FUNCTION_BLOCK "1100_BWTS_CONTROL"   // FB1100, SCL
{ S7_Optimized_Access := 'TRUE' }
VERSION : 0.1
   VAR RETAIN
      State : "SYSTEM_STATES";   // Group of states required for BWT System
      TankData : Array[1..#NumberOfTanks] of "TANK_DATA";   // Group of tank data elements, one per tank on this system
   END_VAR
   VAR
      DECK_MANAGE_START_SUPPLY : "1110_DECK_MANAGE_START_SUPPLY";   // Function to start the deck supply (controlling CV valves 406, 407, 409, 411)
      DECK_MANAGE_STOP_SUPPLY : "1111_DECK_MANAGE_STOP_SUPPLY";   // Function to stop the deck supply (controlling CV valves 406, 407, 409, 411)
   END_VAR
   VAR RETAIN
      GTT_IN : "VALVE_GTT_IN";   // GTT Input data to management block
      GTT_OUT : "VALVE_GTT_OUT";   // GTT Output data from management block
      GTT_Exclusivity : "GTT_EXCLUSIVITY";   // GTT Exclusivity date to manage single valve actuation only
   END_VAR
   VAR
      GTT_MANAGE_VALVES : "1115_GTT_MANAGE_VALVES";
   END_VAR
   VAR RETAIN
      PVVX_IN : "VALVE_PVVX_IN";   // Vent A&B Input data to management blocks
      PVVX_OUT : "VALVE_PVVX_OUT";   // Vent A&B Output data from management blocks
   END_VAR
   VAR
      PVV_MANAGE_VALVES : "1120_PVV_MANAGE_VALVES";
      TANK_CONTROL_FPT : "1105_TANK_CONTROL";   // Tank sub-control block
      TANK_CONTROL_1P : "1105_TANK_CONTROL";   // Tank sub-control block
      TANK_CONTROL_1S : "1105_TANK_CONTROL";   // Tank sub-control block
      TANK_CONTROL_2P : "1105_TANK_CONTROL";   // Tank sub-control block
      TANK_CONTROL_2S : "1105_TANK_CONTROL";   // Tank sub-control block
      TANK_CONTROL_3P : "1105_TANK_CONTROL";   // Tank sub-control block
      TANK_CONTROL_3S : "1105_TANK_CONTROL";   // Tank sub-control block
      TANK_CONTROL_4P : "1105_TANK_CONTROL";   // Tank sub-control block
      TANK_CONTROL_4S : "1105_TANK_CONTROL";   // Tank sub-control block
      TANK_CONTROL_5P : "1105_TANK_CONTROL";   // Tank sub-control block
      TANK_CONTROL_5S : "1105_TANK_CONTROL";   // Tank sub-control block
      TANK_CONTROL_6P : "1105_TANK_CONTROL";   // Tank sub-control block
      TANK_CONTROL_6S : "1105_TANK_CONTROL";   // Tank sub-control block
      TANK_CONTROL_APT : "1105_TANK_CONTROL";   // Tank sub-control block
   END_VAR
   VAR RETAIN
      DWELL_TIMER : TONR_LTIME;   // Dwell Timer to manage Mid-Dwell period
      XEOX_TIMER : TONR_LTIME;   // DeOxygenation and ReOxygenation timer
      XEOX_PAUSE_TIMER : TONR_LTIME;   // The DeOxygenation Pause timer (with retain option)
      XEOX_PausedTime : LTime;   // A counter for the time spent in 'pause' whilst DeOxygenating.
      ShutdownStageReset : Bool := true;   // An reset flag for the shutdown procedure to set the stage to 0 once on a shutdown request.
   END_VAR
   VAR_TEMP
      Index : Int;   // Generic index for for loop parsing
      NextStageCheck : "ALARM_DEMAND_RTN";   // Temporary location for next stage alarm data and stage completion
      NextTreatmentGroup : Int;   // Temporary location for next treatment group calculation
   END_VAR
   VAR CONSTANT
      NumberOfTanks : Int := 14;   // Number of tanks in BWTS
      MaxTimerPT : LTime := LT#106751d;
      State_Init : Int := 0;   // State associated with State.System object.
      State_PreDwell : Int := 1;   // State associated with State.System object.
      State_DeOx : Int := 2;   // State associated with State.System object.
      State_DeOx_SupplyToDeck : Int := 200;   // Sate associated with State.DeOx object.
      State_DeOx_ClosePVV : Int := 201;   // Sate associated with State.DeOx object.
      State_DeOx_OpenGTT : Int := 202;   // Sate associated with State.DeOx object.
      State_DeOx_Monitor : Int := 203;   // Sate associated with State.DeOx object.
      State_DeOx_CloseGTT : Int := 204;   // Sate associated with State.DeOx object.
      State_DeOx_StopSupplyToDeck : Int := 205;   // Sate associated with State.DeOx object.
      State_DwellAndReOx : Int := 3;   // State associated with State.System object.
      State_DwellAndReOx_WaitMidDwell : Int := 300;   // Sate associated with State.ReOx object.
      State_DwellAndReOx_SupplyToDeck : Int := 301;   // Sate associated with State.ReOx object.
      State_DwellAndReOx_OpenPVV : Int := 302;   // Sate associated with State.ReOx object.
      State_DwellAndReOx_OpenGTT : Int := 303;   // Sate associated with State.ReOx object.
      State_DwellAndReOx_Monitor : Int := 304;   // Sate associated with State.ReOx object.
      State_DwellAndReOx_CloseGTT : Int := 305;   // Sate associated with State.ReOx object.
      State_DwellAndReOx_StopSupplyToDeck : Int := 306;   // Sate associated with State.ReOx object.
      State_DwellAndComplete : Int := 4;   // State associated with State.System object.
      State_DwellAndComplete_WaitPostDwell : Int := 400;   // Sate associated with State.Complete object.
      State_DwellAndComplete_Done : Int := 401;   // Sate associated with State.Complete object.
      State_Shutdown : Int := 5;   // State associated with State.System object.
      TankState_Init : Int := 1000;   // State associated with tank sub-control.
      TankState_PreDwell : Int := 1001;   // State associated with tank sub-control.
      TankState_DeOx : Int := 1002;   // State associated with tank sub-control.
      TankState_MidDwell : Int := 1003;   // State associated with tank sub-control.
      TankState_ReOx : Int := 1004;   // State associated with tank sub-control.
      TankState_PostDwell : Int := 1005;   // State associated with tank sub-control.
      TankState_Done : Int := 1006;   // State associated with tank sub-control.
   END_VAR
   // TankData[1].AllocatedTreatmentGroup := 1;
   // TankData[2].AllocatedTreatmentGroup := 1;
   // TankData[3].AllocatedTreatmentGroup := 1;
   // TankData[4].AllocatedTreatmentGroup := 2;
   // TankData[5].AllocatedTreatmentGroup := 2;
   // TankData[6].AllocatedTreatmentGroup := 2;
   // TankData[7].AllocatedTreatmentGroup := 2;
   // TankData[8].AllocatedTreatmentGroup := 3;
   // TankData[9].AllocatedTreatmentGroup := 3;
   // TankData[10].AllocatedTreatmentGroup := 3;
   // TankData[11].AllocatedTreatmentGroup := 4;
   // TankData[12].AllocatedTreatmentGroup := 4;
   // TankData[13].AllocatedTreatmentGroup := 4;
   // TankData[14].AllocatedTreatmentGroup := 4;
   // TankData[1].Active := False;
   // TankData[1].XeOx_Complete := False;
   // TankData[1].Timer_Complete := False;
   // TankData[2].Active := False;
   // TankData[2].XeOx_Complete := False;
   // TankData[2].Timer_Complete := False;
   // TankData[3].Active := False;
   // TankData[3].XeOx_Complete := False;
   // TankData[3].Timer_Complete := False;
   // TankData[4].Active := False;
   // TankData[4].XeOx_Complete := False;
   // TankData[4].Timer_Complete := False;
   // TankData[5].Active := False;
   // TankData[5].XeOx_Complete := False;
   // TankData[5].Timer_Complete := False;
   // TankData[6].Active := False;
   // TankData[6].XeOx_Complete := False;
   // TankData[6].Timer_Complete := False;
   // TankData[7].Active := False;
   // TankData[7].XeOx_Complete := False;
   // TankData[7].Timer_Complete := False;
   // TankData[8].Active := False;
   // TankData[8].XeOx_Complete := False;
   // TankData[8].Timer_Complete := False;
   // TankData[9].Active := False;
   // TankData[9].XeOx_Complete := False;
   // TankData[9].Timer_Complete := False;
   // TankData[10].Active := False;
   // TankData[10].XeOx_Complete := False;
   // TankData[10].Timer_Complete := False;
   // TankData[11].Active := False;
   // TankData[11].XeOx_Complete := False;
   // TankData[11].Timer_Complete := False;
   // TankData[12].Active := False;
   // TankData[12].XeOx_Complete := False;
   // TankData[12].Timer_Complete := False;
   // TankData[13].Active := False;
   // TankData[13].XeOx_Complete := False;
   // TankData[13].Timer_Complete := False;
   // TankData[14].Active := False;
   // TankData[14].XeOx_Complete := False;
   // TankData[14].Timer_Complete := False;
   // DECK_MANAGE_START_SUPPLY.DNC_500CV406.DemandIn := False;
   // DECK_MANAGE_START_SUPPLY.DNC_500CV406.NO_Type := False;
   // DECK_MANAGE_START_SUPPLY.DNC_500CV406.NC_Type := False;
   // DECK_MANAGE_START_SUPPLY.DNC_500CV406.ValveOpenStatus := False;
   // DECK_MANAGE_START_SUPPLY.DNC_500CV406.ValveClsdStatus := False;
   // DECK_MANAGE_START_SUPPLY.DNC_500CV406.DemandOut := False;
   // DECK_MANAGE_START_SUPPLY.DNC_500CV406.DemandComplete := False;
   // DECK_MANAGE_START_SUPPLY.DNC_500CV406.Alarm := False;
   // DECK_MANAGE_START_SUPPLY.DNC_500CV406.Healthy := False;
   // DECK_MANAGE_START_SUPPLY.DNC_500CV406.Config_Error := False;
   // DECK_MANAGE_START_SUPPLY.DNC_500CV406.Sensor_Fault := False;
   // DECK_MANAGE_START_SUPPLY.DNC_500CV406.TRAVEL_TIME.IN := False;
   // DECK_MANAGE_START_SUPPLY.DNC_600CV407.DemandIn := False;
   // DECK_MANAGE_START_SUPPLY.DNC_600CV407.NO_Type := False;
   // DECK_MANAGE_START_SUPPLY.DNC_600CV407.NC_Type := False;
   // DECK_MANAGE_START_SUPPLY.DNC_600CV407.ValveOpenStatus := False;
   // DECK_MANAGE_START_SUPPLY.DNC_600CV407.ValveClsdStatus := False;
   // DECK_MANAGE_START_SUPPLY.DNC_600CV407.DemandOut := False;
   // DECK_MANAGE_START_SUPPLY.DNC_600CV407.DemandComplete := False;
   // DECK_MANAGE_START_SUPPLY.DNC_600CV407.Alarm := False;
   // DECK_MANAGE_START_SUPPLY.DNC_600CV407.Healthy := False;
   // DECK_MANAGE_START_SUPPLY.DNC_600CV407.Config_Error := False;
   // DECK_MANAGE_START_SUPPLY.DNC_600CV407.Sensor_Fault := False;
   // DECK_MANAGE_START_SUPPLY.DNC_600CV407.TRAVEL_TIME.IN := False;
   // DECK_MANAGE_START_SUPPLY.DNC_600CV411.DemandIn := False;
   // DECK_MANAGE_START_SUPPLY.DNC_600CV411.NO_Type := False;
   // DECK_MANAGE_START_SUPPLY.DNC_600CV411.NC_Type := False;
   // DECK_MANAGE_START_SUPPLY.DNC_600CV411.ValveOpenStatus := False;
   // DECK_MANAGE_START_SUPPLY.DNC_600CV411.ValveClsdStatus := False;
   // DECK_MANAGE_START_SUPPLY.DNC_600CV411.DemandOut := False;
   // DECK_MANAGE_START_SUPPLY.DNC_600CV411.DemandComplete := False;
   // DECK_MANAGE_START_SUPPLY.DNC_600CV411.Alarm := False;
   // DECK_MANAGE_START_SUPPLY.DNC_600CV411.Healthy := False;
   // DECK_MANAGE_START_SUPPLY.DNC_600CV411.Config_Error := False;
   // DECK_MANAGE_START_SUPPLY.DNC_600CV411.Sensor_Fault := False;
   // DECK_MANAGE_START_SUPPLY.DNC_600CV411.TRAVEL_TIME.IN := False;
   // DECK_MANAGE_START_SUPPLY.DNC_600CV409.DemandIn := False;
   // DECK_MANAGE_START_SUPPLY.DNC_600CV409.NO_Type := False;
   // DECK_MANAGE_START_SUPPLY.DNC_600CV409.NC_Type := False;
   // DECK_MANAGE_START_SUPPLY.DNC_600CV409.ValveOpenStatus := False;
   // DECK_MANAGE_START_SUPPLY.DNC_600CV409.ValveClsdStatus := False;
   // DECK_MANAGE_START_SUPPLY.DNC_600CV409.DemandOut := False;
   // DECK_MANAGE_START_SUPPLY.DNC_600CV409.DemandComplete := False;
   // DECK_MANAGE_START_SUPPLY.DNC_600CV409.Alarm := False;
   // DECK_MANAGE_START_SUPPLY.DNC_600CV409.Healthy := False;
   // DECK_MANAGE_START_SUPPLY.DNC_600CV409.Config_Error := False;
   // DECK_MANAGE_START_SUPPLY.DNC_600CV409.Sensor_Fault := False;
   // DECK_MANAGE_START_SUPPLY.DNC_600CV409.TRAVEL_TIME.IN := False;
   // DECK_MANAGE_START_SUPPLY.ShutdownDemand := False;
   // DECK_MANAGE_STOP_SUPPLY.DNC_500CV406.DemandIn := False;
   // DECK_MANAGE_STOP_SUPPLY.DNC_500CV406.NO_Type := False;
   // DECK_MANAGE_STOP_SUPPLY.DNC_500CV406.NC_Type := False;
   // DECK_MANAGE_STOP_SUPPLY.DNC_500CV406.ValveOpenStatus := False;
   // DECK_MANAGE_STOP_SUPPLY.DNC_500CV406.ValveClsdStatus := False;
   // DECK_MANAGE_STOP_SUPPLY.DNC_500CV406.DemandOut := False;
   // DECK_MANAGE_STOP_SUPPLY.DNC_500CV406.DemandComplete := False;
   // DECK_MANAGE_STOP_SUPPLY.DNC_500CV406.Alarm := False;
   // DECK_MANAGE_STOP_SUPPLY.DNC_500CV406.Healthy := False;
   // DECK_MANAGE_STOP_SUPPLY.DNC_500CV406.Config_Error := False;
   // DECK_MANAGE_STOP_SUPPLY.DNC_500CV406.Sensor_Fault := False;
   // DECK_MANAGE_STOP_SUPPLY.DNC_500CV406.TRAVEL_TIME.IN := False;
   // DECK_MANAGE_STOP_SUPPLY.DNC_600CV407.DemandIn := False;
   // DECK_MANAGE_STOP_SUPPLY.DNC_600CV407.NO_Type := False;
   // DECK_MANAGE_STOP_SUPPLY.DNC_600CV407.NC_Type := False;
   // DECK_MANAGE_STOP_SUPPLY.DNC_600CV407.ValveOpenStatus := False;
   // DECK_MANAGE_STOP_SUPPLY.DNC_600CV407.ValveClsdStatus := False;
   // DECK_MANAGE_STOP_SUPPLY.DNC_600CV407.DemandOut := False;
   // DECK_MANAGE_STOP_SUPPLY.DNC_600CV407.DemandComplete := False;
   // DECK_MANAGE_STOP_SUPPLY.DNC_600CV407.Alarm := False;
   // DECK_MANAGE_STOP_SUPPLY.DNC_600CV407.Healthy := False;
   // DECK_MANAGE_STOP_SUPPLY.DNC_600CV407.Config_Error := False;
   // DECK_MANAGE_STOP_SUPPLY.DNC_600CV407.Sensor_Fault := False;
   // DECK_MANAGE_STOP_SUPPLY.DNC_600CV407.TRAVEL_TIME.IN := False;
   // DECK_MANAGE_STOP_SUPPLY.DNC_600CV411.DemandIn := False;
   // DECK_MANAGE_STOP_SUPPLY.DNC_600CV411.NO_Type := False;
   // DECK_MANAGE_STOP_SUPPLY.DNC_600CV411.NC_Type := False;
   // DECK_MANAGE_STOP_SUPPLY.DNC_600CV411.ValveOpenStatus := False;
   // DECK_MANAGE_STOP_SUPPLY.DNC_600CV411.ValveClsdStatus := False;
   // DECK_MANAGE_STOP_SUPPLY.DNC_600CV411.DemandOut := False;
   // DECK_MANAGE_STOP_SUPPLY.DNC_600CV411.DemandComplete := False;
   // DECK_MANAGE_STOP_SUPPLY.DNC_600CV411.Alarm := False;
   // DECK_MANAGE_STOP_SUPPLY.DNC_600CV411.Healthy := False;
   // DECK_MANAGE_STOP_SUPPLY.DNC_600CV411.Config_Error := False;
   // DECK_MANAGE_STOP_SUPPLY.DNC_600CV411.Sensor_Fault := False;
   // DECK_MANAGE_STOP_SUPPLY.DNC_600CV411.TRAVEL_TIME.IN := False;
   // DECK_MANAGE_STOP_SUPPLY.DNC_600CV409.DemandIn := False;
   // DECK_MANAGE_STOP_SUPPLY.DNC_600CV409.NO_Type := False;
   // DECK_MANAGE_STOP_SUPPLY.DNC_600CV409.NC_Type := False;
   // DECK_MANAGE_STOP_SUPPLY.DNC_600CV409.ValveOpenStatus := False;
   // DECK_MANAGE_STOP_SUPPLY.DNC_600CV409.ValveClsdStatus := False;
   // DECK_MANAGE_STOP_SUPPLY.DNC_600CV409.DemandOut := False;
   // DECK_MANAGE_STOP_SUPPLY.DNC_600CV409.DemandComplete := False;
   // DECK_MANAGE_STOP_SUPPLY.DNC_600CV409.Alarm := False;
   // DECK_MANAGE_STOP_SUPPLY.DNC_600CV409.Healthy := False;
   // DECK_MANAGE_STOP_SUPPLY.DNC_600CV409.Config_Error := False;
   // DECK_MANAGE_STOP_SUPPLY.DNC_600CV409.Sensor_Fault := False;
   // DECK_MANAGE_STOP_SUPPLY.DNC_600CV409.TRAVEL_TIME.IN := False;
   // DECK_MANAGE_STOP_SUPPLY.TON_DELAY.IN := False;
   // DECK_MANAGE_STOP_SUPPLY.ShutdownDemand := False;
   // DECK_MANAGE_STOP_SUPPLY.StopDeckSupplyDone := False;
   // GTT_IN.GTT_Actuate[1] := False;
   // GTT_IN.GTT_Actuate[2] := False;
   // GTT_IN.GTT_Actuate[3] := False;
   // GTT_IN.GTT_Actuate[4] := False;
   // GTT_IN.GTT_Actuate[5] := False;
   // GTT_IN.GTT_Actuate[6] := False;
   // GTT_IN.GTT_Actuate[7] := False;
   // GTT_IN.GTT_Actuate[8] := False;
   // GTT_IN.GTT_Actuate[9] := False;
   // GTT_IN.GTT_Actuate[10] := False;
   // GTT_IN.GTT_Actuate[11] := False;
   // GTT_IN.GTT_Actuate[12] := False;
   // GTT_IN.GTT_Actuate[13] := False;
   // GTT_IN.GTT_Actuate[14] := False;
   // GTT_IN.GTT_ValveDemands[1] := False;
   // GTT_IN.GTT_ValveDemands[2] := False;
   // GTT_IN.GTT_ValveDemands[3] := False;
   // GTT_IN.GTT_ValveDemands[4] := False;
   // GTT_IN.GTT_ValveDemands[5] := False;
   // GTT_IN.GTT_ValveDemands[6] := False;
   // GTT_IN.GTT_ValveDemands[7] := False;
   // GTT_IN.GTT_ValveDemands[8] := False;
   // GTT_IN.GTT_ValveDemands[9] := False;
   // GTT_IN.GTT_ValveDemands[10] := False;
   // GTT_IN.GTT_ValveDemands[11] := False;
   // GTT_IN.GTT_ValveDemands[12] := False;
   // GTT_IN.GTT_ValveDemands[13] := False;
   // GTT_IN.GTT_ValveDemands[14] := False;
   // GTT_OUT.GTT_DemandsCompleted[1] := False;
   // GTT_OUT.GTT_DemandsCompleted[2] := False;
   // GTT_OUT.GTT_DemandsCompleted[3] := False;
   // GTT_OUT.GTT_DemandsCompleted[4] := False;
   // GTT_OUT.GTT_DemandsCompleted[5] := False;
   // GTT_OUT.GTT_DemandsCompleted[6] := False;
   // GTT_OUT.GTT_DemandsCompleted[7] := False;
   // GTT_OUT.GTT_DemandsCompleted[8] := False;
   // GTT_OUT.GTT_DemandsCompleted[9] := False;
   // GTT_OUT.GTT_DemandsCompleted[10] := False;
   // GTT_OUT.GTT_DemandsCompleted[11] := False;
   // GTT_OUT.GTT_DemandsCompleted[12] := False;
   // GTT_OUT.GTT_DemandsCompleted[13] := False;
   // GTT_OUT.GTT_DemandsCompleted[14] := False;
   // GTT_OUT.GTT_Alarms[1] := False;
   // GTT_OUT.GTT_Alarms[2] := False;
   // GTT_OUT.GTT_Alarms[3] := False;
   // GTT_OUT.GTT_Alarms[4] := False;
   // GTT_OUT.GTT_Alarms[5] := False;
   // GTT_OUT.GTT_Alarms[6] := False;
   // GTT_OUT.GTT_Alarms[7] := False;
   // GTT_OUT.GTT_Alarms[8] := False;
   // GTT_OUT.GTT_Alarms[9] := False;
   // GTT_OUT.GTT_Alarms[10] := False;
   // GTT_OUT.GTT_Alarms[11] := False;
   // GTT_OUT.GTT_Alarms[12] := False;
   // GTT_OUT.GTT_Alarms[13] := False;
   // GTT_OUT.GTT_Alarms[14] := False;
   // GTT_Exclusivity.Tank_Exclusivity := False;
   // GTT_MANAGE_VALVES.GTT_IN.GTT_Actuate[1] := False;
   // GTT_MANAGE_VALVES.GTT_IN.GTT_Actuate[2] := False;
   // GTT_MANAGE_VALVES.GTT_IN.GTT_Actuate[3] := False;
   // GTT_MANAGE_VALVES.GTT_IN.GTT_Actuate[4] := False;
   // GTT_MANAGE_VALVES.GTT_IN.GTT_Actuate[5] := False;
   // GTT_MANAGE_VALVES.GTT_IN.GTT_Actuate[6] := False;
   // GTT_MANAGE_VALVES.GTT_IN.GTT_Actuate[7] := False;
   // GTT_MANAGE_VALVES.GTT_IN.GTT_Actuate[8] := False;
   // GTT_MANAGE_VALVES.GTT_IN.GTT_Actuate[9] := False;
   // GTT_MANAGE_VALVES.GTT_IN.GTT_Actuate[10] := False;
   // GTT_MANAGE_VALVES.GTT_IN.GTT_Actuate[11] := False;
   // GTT_MANAGE_VALVES.GTT_IN.GTT_Actuate[12] := False;
   // GTT_MANAGE_VALVES.GTT_IN.GTT_Actuate[13] := False;
   // GTT_MANAGE_VALVES.GTT_IN.GTT_Actuate[14] := False;
   // GTT_MANAGE_VALVES.GTT_IN.GTT_ValveDemands[1] := False;
   // GTT_MANAGE_VALVES.GTT_IN.GTT_ValveDemands[2] := False;
   // GTT_MANAGE_VALVES.GTT_IN.GTT_ValveDemands[3] := False;
   // GTT_MANAGE_VALVES.GTT_IN.GTT_ValveDemands[4] := False;
   // GTT_MANAGE_VALVES.GTT_IN.GTT_ValveDemands[5] := False;
   // GTT_MANAGE_VALVES.GTT_IN.GTT_ValveDemands[6] := False;
   // GTT_MANAGE_VALVES.GTT_IN.GTT_ValveDemands[7] := False;
   // GTT_MANAGE_VALVES.GTT_IN.GTT_ValveDemands[8] := False;
   // GTT_MANAGE_VALVES.GTT_IN.GTT_ValveDemands[9] := False;
   // GTT_MANAGE_VALVES.GTT_IN.GTT_ValveDemands[10] := False;
   // GTT_MANAGE_VALVES.GTT_IN.GTT_ValveDemands[11] := False;
   // GTT_MANAGE_VALVES.GTT_IN.GTT_ValveDemands[12] := False;
   // GTT_MANAGE_VALVES.GTT_IN.GTT_ValveDemands[13] := False;
   // GTT_MANAGE_VALVES.GTT_IN.GTT_ValveDemands[14] := False;
   // GTT_MANAGE_VALVES.DNC_FPT_GTT.DemandIn := False;
   // GTT_MANAGE_VALVES.DNC_FPT_GTT.NO_Type := False;
   // GTT_MANAGE_VALVES.DNC_FPT_GTT.NC_Type := False;
   // GTT_MANAGE_VALVES.DNC_FPT_GTT.ValveOpenStatus := False;
   // GTT_MANAGE_VALVES.DNC_FPT_GTT.ValveClsdStatus := False;
   // GTT_MANAGE_VALVES.DNC_FPT_GTT.DemandOut := False;
   // GTT_MANAGE_VALVES.DNC_FPT_GTT.DemandComplete := False;
   // GTT_MANAGE_VALVES.DNC_FPT_GTT.Alarm := False;
   // GTT_MANAGE_VALVES.DNC_FPT_GTT.Healthy := False;
   // GTT_MANAGE_VALVES.DNC_FPT_GTT.Config_Error := False;
   // GTT_MANAGE_VALVES.DNC_FPT_GTT.Sensor_Fault := False;
   // GTT_MANAGE_VALVES.DNC_FPT_GTT.TRAVEL_TIME.IN := False;
   // GTT_MANAGE_VALVES.DNC_1P_GTT.DemandIn := False;
   // GTT_MANAGE_VALVES.DNC_1P_GTT.NO_Type := False;
   // GTT_MANAGE_VALVES.DNC_1P_GTT.NC_Type := False;
   // GTT_MANAGE_VALVES.DNC_1P_GTT.ValveOpenStatus := False;
   // GTT_MANAGE_VALVES.DNC_1P_GTT.ValveClsdStatus := False;
   // GTT_MANAGE_VALVES.DNC_1P_GTT.DemandOut := False;
   // GTT_MANAGE_VALVES.DNC_1P_GTT.DemandComplete := False;
   // GTT_MANAGE_VALVES.DNC_1P_GTT.Alarm := False;
   // GTT_MANAGE_VALVES.DNC_1P_GTT.Healthy := False;
   // GTT_MANAGE_VALVES.DNC_1P_GTT.Config_Error := False;
   // GTT_MANAGE_VALVES.DNC_1P_GTT.Sensor_Fault := False;
   // GTT_MANAGE_VALVES.DNC_1P_GTT.TRAVEL_TIME.IN := False;
   // GTT_MANAGE_VALVES.DNC_1S_GTT.DemandIn := False;
   // GTT_MANAGE_VALVES.DNC_1S_GTT.NO_Type := False;
   // GTT_MANAGE_VALVES.DNC_1S_GTT.NC_Type := False;
   // GTT_MANAGE_VALVES.DNC_1S_GTT.ValveOpenStatus := False;
   // GTT_MANAGE_VALVES.DNC_1S_GTT.ValveClsdStatus := False;
   // GTT_MANAGE_VALVES.DNC_1S_GTT.DemandOut := False;
   // GTT_MANAGE_VALVES.DNC_1S_GTT.DemandComplete := False;
   // GTT_MANAGE_VALVES.DNC_1S_GTT.Alarm := False;
   // GTT_MANAGE_VALVES.DNC_1S_GTT.Healthy := False;
   // GTT_MANAGE_VALVES.DNC_1S_GTT.Config_Error := False;
   // GTT_MANAGE_VALVES.DNC_1S_GTT.Sensor_Fault := False;
   // GTT_MANAGE_VALVES.DNC_1S_GTT.TRAVEL_TIME.IN := False;
   // GTT_MANAGE_VALVES.DNC_2P_GTT.DemandIn := False;
   // GTT_MANAGE_VALVES.DNC_2P_GTT.NO_Type := False;
   // GTT_MANAGE_VALVES.DNC_2P_GTT.NC_Type := False;
   // GTT_MANAGE_VALVES.DNC_2P_GTT.ValveOpenStatus := False;
   // GTT_MANAGE_VALVES.DNC_2P_GTT.ValveClsdStatus := False;
   // GTT_MANAGE_VALVES.DNC_2P_GTT.DemandOut := False;
   // GTT_MANAGE_VALVES.DNC_2P_GTT.DemandComplete := False;
   // GTT_MANAGE_VALVES.DNC_2P_GTT.Alarm := False;
   // GTT_MANAGE_VALVES.DNC_2P_GTT.Healthy := False;
   // GTT_MANAGE_VALVES.DNC_2P_GTT.Config_Error := False;
   // GTT_MANAGE_VALVES.DNC_2P_GTT.Sensor_Fault := False;
   // GTT_MANAGE_VALVES.DNC_2P_GTT.TRAVEL_TIME.IN := False;
   // GTT_MANAGE_VALVES.DNC_2S_GTT.DemandIn := False;
   // GTT_MANAGE_VALVES.DNC_2S_GTT.NO_Type := False;
   // GTT_MANAGE_VALVES.DNC_2S_GTT.NC_Type := False;
   // GTT_MANAGE_VALVES.DNC_2S_GTT.ValveOpenStatus := False;
   // GTT_MANAGE_VALVES.DNC_2S_GTT.ValveClsdStatus := False;
   // GTT_MANAGE_VALVES.DNC_2S_GTT.DemandOut := False;
   // GTT_MANAGE_VALVES.DNC_2S_GTT.DemandComplete := False;
   // GTT_MANAGE_VALVES.DNC_2S_GTT.Alarm := False;
   // GTT_MANAGE_VALVES.DNC_2S_GTT.Healthy := False;
   // GTT_MANAGE_VALVES.DNC_2S_GTT.Config_Error := False;
   // GTT_MANAGE_VALVES.DNC_2S_GTT.Sensor_Fault := False;
   // GTT_MANAGE_VALVES.DNC_2S_GTT.TRAVEL_TIME.IN := False;
   // GTT_MANAGE_VALVES.DNC_3P_GTT.DemandIn := False;
   // GTT_MANAGE_VALVES.DNC_3P_GTT.NO_Type := False;
   // GTT_MANAGE_VALVES.DNC_3P_GTT.NC_Type := False;
   // GTT_MANAGE_VALVES.DNC_3P_GTT.ValveOpenStatus := False;
   // GTT_MANAGE_VALVES.DNC_3P_GTT.ValveClsdStatus := False;
   // GTT_MANAGE_VALVES.DNC_3P_GTT.DemandOut := False;
   // GTT_MANAGE_VALVES.DNC_3P_GTT.DemandComplete := False;
   // GTT_MANAGE_VALVES.DNC_3P_GTT.Alarm := False;
   // GTT_MANAGE_VALVES.DNC_3P_GTT.Healthy := False;
   // GTT_MANAGE_VALVES.DNC_3P_GTT.Config_Error := False;
   // GTT_MANAGE_VALVES.DNC_3P_GTT.Sensor_Fault := False;
   // GTT_MANAGE_VALVES.DNC_3P_GTT.TRAVEL_TIME.IN := False;
   // GTT_MANAGE_VALVES.DNC_3S_GTT.DemandIn := False;
   // GTT_MANAGE_VALVES.DNC_3S_GTT.NO_Type := False;
   // GTT_MANAGE_VALVES.DNC_3S_GTT.NC_Type := False;
   // GTT_MANAGE_VALVES.DNC_3S_GTT.ValveOpenStatus := False;
   // GTT_MANAGE_VALVES.DNC_3S_GTT.ValveClsdStatus := False;
   // GTT_MANAGE_VALVES.DNC_3S_GTT.DemandOut := False;
   // GTT_MANAGE_VALVES.DNC_3S_GTT.DemandComplete := False;
   // GTT_MANAGE_VALVES.DNC_3S_GTT.Alarm := False;
   // GTT_MANAGE_VALVES.DNC_3S_GTT.Healthy := False;
   // GTT_MANAGE_VALVES.DNC_3S_GTT.Config_Error := False;
   // GTT_MANAGE_VALVES.DNC_3S_GTT.Sensor_Fault := False;
   // GTT_MANAGE_VALVES.DNC_3S_GTT.TRAVEL_TIME.IN := False;
   // GTT_MANAGE_VALVES.DNC_4P_GTT.DemandIn := False;
   // GTT_MANAGE_VALVES.DNC_4P_GTT.NO_Type := False;
   // GTT_MANAGE_VALVES.DNC_4P_GTT.NC_Type := False;
   // GTT_MANAGE_VALVES.DNC_4P_GTT.ValveOpenStatus := False;
   // GTT_MANAGE_VALVES.DNC_4P_GTT.ValveClsdStatus := False;
   // GTT_MANAGE_VALVES.DNC_4P_GTT.DemandOut := False;
   // GTT_MANAGE_VALVES.DNC_4P_GTT.DemandComplete := False;
   // GTT_MANAGE_VALVES.DNC_4P_GTT.Alarm := False;
   // GTT_MANAGE_VALVES.DNC_4P_GTT.Healthy := False;
   // GTT_MANAGE_VALVES.DNC_4P_GTT.Config_Error := False;
   // GTT_MANAGE_VALVES.DNC_4P_GTT.Sensor_Fault := False;
   // GTT_MANAGE_VALVES.DNC_4P_GTT.TRAVEL_TIME.IN := False;
   // GTT_MANAGE_VALVES.DNC_4S_GTT.DemandIn := False;
   // GTT_MANAGE_VALVES.DNC_4S_GTT.NO_Type := False;
   // GTT_MANAGE_VALVES.DNC_4S_GTT.NC_Type := False;
   // GTT_MANAGE_VALVES.DNC_4S_GTT.ValveOpenStatus := False;
   // GTT_MANAGE_VALVES.DNC_4S_GTT.ValveClsdStatus := False;
   // GTT_MANAGE_VALVES.DNC_4S_GTT.DemandOut := False;
   // GTT_MANAGE_VALVES.DNC_4S_GTT.DemandComplete := False;
   // GTT_MANAGE_VALVES.DNC_4S_GTT.Alarm := False;
   // GTT_MANAGE_VALVES.DNC_4S_GTT.Healthy := False;
   // GTT_MANAGE_VALVES.DNC_4S_GTT.Config_Error := False;
   // GTT_MANAGE_VALVES.DNC_4S_GTT.Sensor_Fault := False;
   // GTT_MANAGE_VALVES.DNC_4S_GTT.TRAVEL_TIME.IN := False;
   // GTT_MANAGE_VALVES.DNC_5P_GTT.DemandIn := False;
   // GTT_MANAGE_VALVES.DNC_5P_GTT.NO_Type := False;
   // GTT_MANAGE_VALVES.DNC_5P_GTT.NC_Type := False;
   // GTT_MANAGE_VALVES.DNC_5P_GTT.ValveOpenStatus := False;
   // GTT_MANAGE_VALVES.DNC_5P_GTT.ValveClsdStatus := False;
   // GTT_MANAGE_VALVES.DNC_5P_GTT.DemandOut := False;
   // GTT_MANAGE_VALVES.DNC_5P_GTT.DemandComplete := False;
   // GTT_MANAGE_VALVES.DNC_5P_GTT.Alarm := False;
   // GTT_MANAGE_VALVES.DNC_5P_GTT.Healthy := False;
   // GTT_MANAGE_VALVES.DNC_5P_GTT.Config_Error := False;
   // GTT_MANAGE_VALVES.DNC_5P_GTT.Sensor_Fault := False;
   // GTT_MANAGE_VALVES.DNC_5P_GTT.TRAVEL_TIME.IN := False;
   // GTT_MANAGE_VALVES.DNC_5S_GTT.DemandIn := False;
   // GTT_MANAGE_VALVES.DNC_5S_GTT.NO_Type := False;
   // GTT_MANAGE_VALVES.DNC_5S_GTT.NC_Type := False;
   // GTT_MANAGE_VALVES.DNC_5S_GTT.ValveOpenStatus := False;
   // GTT_MANAGE_VALVES.DNC_5S_GTT.ValveClsdStatus := False;
   // GTT_MANAGE_VALVES.DNC_5S_GTT.DemandOut := False;
   // GTT_MANAGE_VALVES.DNC_5S_GTT.DemandComplete := False;
   // GTT_MANAGE_VALVES.DNC_5S_GTT.Alarm := False;
   // GTT_MANAGE_VALVES.DNC_5S_GTT.Healthy := False;
   // GTT_MANAGE_VALVES.DNC_5S_GTT.Config_Error := False;
   // GTT_MANAGE_VALVES.DNC_5S_GTT.Sensor_Fault := False;
   // GTT_MANAGE_VALVES.DNC_5S_GTT.TRAVEL_TIME.IN := False;
   // GTT_MANAGE_VALVES.DNC_6P_GTT.DemandIn := False;
   // GTT_MANAGE_VALVES.DNC_6P_GTT.NO_Type := False;
   // GTT_MANAGE_VALVES.DNC_6P_GTT.NC_Type := False;
   // GTT_MANAGE_VALVES.DNC_6P_GTT.ValveOpenStatus := False;
   // GTT_MANAGE_VALVES.DNC_6P_GTT.ValveClsdStatus := False;
   // GTT_MANAGE_VALVES.DNC_6P_GTT.DemandOut := False;
   // GTT_MANAGE_VALVES.DNC_6P_GTT.DemandComplete := False;
   // GTT_MANAGE_VALVES.DNC_6P_GTT.Alarm := False;
   // GTT_MANAGE_VALVES.DNC_6P_GTT.Healthy := False;
   // GTT_MANAGE_VALVES.DNC_6P_GTT.Config_Error := False;
   // GTT_MANAGE_VALVES.DNC_6P_GTT.Sensor_Fault := False;
   // GTT_MANAGE_VALVES.DNC_6P_GTT.TRAVEL_TIME.IN := False;
   // GTT_MANAGE_VALVES.DNC_6S_GTT.DemandIn := False;
   // GTT_MANAGE_VALVES.DNC_6S_GTT.NO_Type := False;
   // GTT_MANAGE_VALVES.DNC_6S_GTT.NC_Type := False;
   // GTT_MANAGE_VALVES.DNC_6S_GTT.ValveOpenStatus := False;
   // GTT_MANAGE_VALVES.DNC_6S_GTT.ValveClsdStatus := False;
   // GTT_MANAGE_VALVES.DNC_6S_GTT.DemandOut := False;
   // GTT_MANAGE_VALVES.DNC_6S_GTT.DemandComplete := False;
   // GTT_MANAGE_VALVES.DNC_6S_GTT.Alarm := False;
   // GTT_MANAGE_VALVES.DNC_6S_GTT.Healthy := False;
   // GTT_MANAGE_VALVES.DNC_6S_GTT.Config_Error := False;
   // GTT_MANAGE_VALVES.DNC_6S_GTT.Sensor_Fault := False;
   // GTT_MANAGE_VALVES.DNC_6S_GTT.TRAVEL_TIME.IN := False;
   // GTT_MANAGE_VALVES.DNC_APT_GTT.DemandIn := False;
   // GTT_MANAGE_VALVES.DNC_APT_GTT.NO_Type := False;
   // GTT_MANAGE_VALVES.DNC_APT_GTT.NC_Type := False;
   // GTT_MANAGE_VALVES.DNC_APT_GTT.ValveOpenStatus := False;
   // GTT_MANAGE_VALVES.DNC_APT_GTT.ValveClsdStatus := False;
   // GTT_MANAGE_VALVES.DNC_APT_GTT.DemandOut := False;
   // GTT_MANAGE_VALVES.DNC_APT_GTT.DemandComplete := False;
   // GTT_MANAGE_VALVES.DNC_APT_GTT.Alarm := False;
   // GTT_MANAGE_VALVES.DNC_APT_GTT.Healthy := False;
   // GTT_MANAGE_VALVES.DNC_APT_GTT.Config_Error := False;
   // GTT_MANAGE_VALVES.DNC_APT_GTT.Sensor_Fault := False;
   // GTT_MANAGE_VALVES.DNC_APT_GTT.TRAVEL_TIME.IN := False;
   // PVVX_IN.PVVx_Actuate[1] := False;
   // PVVX_IN.PVVx_Actuate[2] := False;
   // PVVX_IN.PVVx_Actuate[3] := False;
   // PVVX_IN.PVVx_Actuate[4] := False;
   // PVVX_IN.PVVx_Actuate[5] := False;
   // PVVX_IN.PVVx_Actuate[6] := False;
   // PVVX_IN.PVVx_Actuate[7] := False;
   // PVVX_IN.PVVx_Actuate[8] := False;
   // PVVX_IN.PVVx_Actuate[9] := False;
   // PVVX_IN.PVVx_Actuate[10] := False;
   // PVVX_IN.PVVx_Actuate[11] := False;
   // PVVX_IN.PVVx_Actuate[12] := False;
   // PVVX_IN.PVVx_Actuate[13] := False;
   // PVVX_IN.PVVx_Actuate[14] := False;
   // PVVX_IN.PVVA_ValveDemands[1] := False;
   // PVVX_IN.PVVA_ValveDemands[2] := False;
   // PVVX_IN.PVVA_ValveDemands[3] := False;
   // PVVX_IN.PVVA_ValveDemands[4] := False;
   // PVVX_IN.PVVA_ValveDemands[5] := False;
   // PVVX_IN.PVVA_ValveDemands[6] := False;
   // PVVX_IN.PVVA_ValveDemands[7] := False;
   // PVVX_IN.PVVA_ValveDemands[8] := False;
   // PVVX_IN.PVVA_ValveDemands[9] := False;
   // PVVX_IN.PVVA_ValveDemands[10] := False;
   // PVVX_IN.PVVA_ValveDemands[11] := False;
   // PVVX_IN.PVVA_ValveDemands[12] := False;
   // PVVX_IN.PVVA_ValveDemands[13] := False;
   // PVVX_IN.PVVA_ValveDemands[14] := False;
   // PVVX_IN.PVVB_ValveDemands[1] := False;
   // PVVX_IN.PVVB_ValveDemands[2] := False;
   // PVVX_IN.PVVB_ValveDemands[3] := False;
   // PVVX_IN.PVVB_ValveDemands[4] := False;
   // PVVX_IN.PVVB_ValveDemands[5] := False;
   // PVVX_IN.PVVB_ValveDemands[6] := False;
   // PVVX_IN.PVVB_ValveDemands[7] := False;
   // PVVX_IN.PVVB_ValveDemands[8] := False;
   // PVVX_IN.PVVB_ValveDemands[9] := False;
   // PVVX_IN.PVVB_ValveDemands[10] := False;
   // PVVX_IN.PVVB_ValveDemands[11] := False;
   // PVVX_IN.PVVB_ValveDemands[12] := False;
   // PVVX_IN.PVVB_ValveDemands[13] := False;
   // PVVX_IN.PVVB_ValveDemands[14] := False;
   // PVVX_OUT.PVVA_DemandsCompleted[1] := False;
   // PVVX_OUT.PVVA_DemandsCompleted[2] := False;
   // PVVX_OUT.PVVA_DemandsCompleted[3] := False;
   // PVVX_OUT.PVVA_DemandsCompleted[4] := False;
   // PVVX_OUT.PVVA_DemandsCompleted[5] := False;
   // PVVX_OUT.PVVA_DemandsCompleted[6] := False;
   // PVVX_OUT.PVVA_DemandsCompleted[7] := False;
   // PVVX_OUT.PVVA_DemandsCompleted[8] := False;
   // PVVX_OUT.PVVA_DemandsCompleted[9] := False;
   // PVVX_OUT.PVVA_DemandsCompleted[10] := False;
   // PVVX_OUT.PVVA_DemandsCompleted[11] := False;
   // PVVX_OUT.PVVA_DemandsCompleted[12] := False;
   // PVVX_OUT.PVVA_DemandsCompleted[13] := False;
   // PVVX_OUT.PVVA_DemandsCompleted[14] := False;
   // PVVX_OUT.PVVA_Alarms[1] := False;
   // PVVX_OUT.PVVA_Alarms[2] := False;
   // PVVX_OUT.PVVA_Alarms[3] := False;
   // PVVX_OUT.PVVA_Alarms[4] := False;
   // PVVX_OUT.PVVA_Alarms[5] := False;
   // PVVX_OUT.PVVA_Alarms[6] := False;
   // PVVX_OUT.PVVA_Alarms[7] := False;
   // PVVX_OUT.PVVA_Alarms[8] := False;
   // PVVX_OUT.PVVA_Alarms[9] := False;
   // PVVX_OUT.PVVA_Alarms[10] := False;
   // PVVX_OUT.PVVA_Alarms[11] := False;
   // PVVX_OUT.PVVA_Alarms[12] := False;
   // PVVX_OUT.PVVA_Alarms[13] := False;
   // PVVX_OUT.PVVA_Alarms[14] := False;
   // PVVX_OUT.PVVB_DemandsCompleted[1] := False;
   // PVVX_OUT.PVVB_DemandsCompleted[2] := False;
   // PVVX_OUT.PVVB_DemandsCompleted[3] := False;
   // PVVX_OUT.PVVB_DemandsCompleted[4] := False;
   // PVVX_OUT.PVVB_DemandsCompleted[5] := False;
   // PVVX_OUT.PVVB_DemandsCompleted[6] := False;
   // PVVX_OUT.PVVB_DemandsCompleted[7] := False;
   // PVVX_OUT.PVVB_DemandsCompleted[8] := False;
   // PVVX_OUT.PVVB_DemandsCompleted[9] := False;
   // PVVX_OUT.PVVB_DemandsCompleted[10] := False;
   // PVVX_OUT.PVVB_DemandsCompleted[11] := False;
   // PVVX_OUT.PVVB_DemandsCompleted[12] := False;
   // PVVX_OUT.PVVB_DemandsCompleted[13] := False;
   // PVVX_OUT.PVVB_DemandsCompleted[14] := False;
   // PVVX_OUT.PVVB_Alarms[1] := False;
   // PVVX_OUT.PVVB_Alarms[2] := False;
   // PVVX_OUT.PVVB_Alarms[3] := False;
   // PVVX_OUT.PVVB_Alarms[4] := False;
   // PVVX_OUT.PVVB_Alarms[5] := False;
   // PVVX_OUT.PVVB_Alarms[6] := False;
   // PVVX_OUT.PVVB_Alarms[7] := False;
   // PVVX_OUT.PVVB_Alarms[8] := False;
   // PVVX_OUT.PVVB_Alarms[9] := False;
   // PVVX_OUT.PVVB_Alarms[10] := False;
   // PVVX_OUT.PVVB_Alarms[11] := False;
   // PVVX_OUT.PVVB_Alarms[12] := False;
   // PVVX_OUT.PVVB_Alarms[13] := False;
   // PVVX_OUT.PVVB_Alarms[14] := False;
   // PVV_MANAGE_VALVES.PVVX_IN.PVVx_Actuate[1] := False;
   // PVV_MANAGE_VALVES.PVVX_IN.PVVx_Actuate[2] := False;
   // PVV_MANAGE_VALVES.PVVX_IN.PVVx_Actuate[3] := False;
   // PVV_MANAGE_VALVES.PVVX_IN.PVVx_Actuate[4] := False;
   // PVV_MANAGE_VALVES.PVVX_IN.PVVx_Actuate[5] := False;
   // PVV_MANAGE_VALVES.PVVX_IN.PVVx_Actuate[6] := False;
   // PVV_MANAGE_VALVES.PVVX_IN.PVVx_Actuate[7] := False;
   // PVV_MANAGE_VALVES.PVVX_IN.PVVx_Actuate[8] := False;
   // PVV_MANAGE_VALVES.PVVX_IN.PVVx_Actuate[9] := False;
   // PVV_MANAGE_VALVES.PVVX_IN.PVVx_Actuate[10] := False;
   // PVV_MANAGE_VALVES.PVVX_IN.PVVx_Actuate[11] := False;
   // PVV_MANAGE_VALVES.PVVX_IN.PVVx_Actuate[12] := False;
   // PVV_MANAGE_VALVES.PVVX_IN.PVVx_Actuate[13] := False;
   // PVV_MANAGE_VALVES.PVVX_IN.PVVx_Actuate[14] := False;
   // PVV_MANAGE_VALVES.PVVX_IN.PVVA_ValveDemands[1] := False;
   // PVV_MANAGE_VALVES.PVVX_IN.PVVA_ValveDemands[2] := False;